screen "SP" 800x480, template "Main"
   GraphicView "Graphic view_1" at 20,61 size 347x209; Picture "clean2"
   TextField "Text field_1" at 288,5 size 156x47; Text 'Уставки'
   TextField "Text field_2" at 138,75 size 112x33; Text 'Дозация'
   TextField "Text field_12" at 28,137 size 34x23; Text 'С ='
   TextField "Text field_13" at 132,138 size 67x23; Text '% масс'
   GraphicView "Graphic view_2" at 64,133 size 66x33; Picture "input_1"
   IOField "I/O field_1" at 68,136 size 58x27; Authorization "Operator"; FormatPattern 9.99
      ProcessValue <- "Logick_DB_SP"
   GraphicView "Graphic view_5" at 368,61 size 347x209; Picture "clean2"
   TextField "Text field_21" at 436,75 size 211x33; Text 'Перемешивание'
   TextField "Text field_22" at 381,129 size 215x23; Text 'Первое перемешивание:'
   TextField "Text field_23" at 667,129 size 17x23; Text 'м'
   GraphicView "Graphic view_6" at 599,124 size 66x33; Picture "input_1"
   IOField "I/O field_3" at 603,127 size 58x27; Authorization "Operator"; FormatPattern 99
      ProcessValue <- "Logick_DB_T_M_SP_M"
   GraphicView "Graphic view_8" at 21,270 size 347x209; Picture "clean2"
   TextField "Text field_14" at 108,283 size 174x33; Text 'Реле протока'
      Visibility <- "CONFIG_Config_Use_DL"
   GraphicView "Graphic view_11" at 368,270 size 347x209; Picture "clean2"
   TextField "Text field_9" at 430,284 size 223x33; Text 'Контроль уровня'
   TextField "Text field_3" at 76,118 size 43x17; Text 'макс 1'
   TextField "Text field_4" at 71,163 size 53x17; Text 'мин 0.05'
   TextField "Text field_5" at 29,177 size 192x23; Text 'Литров на 1 дозацию:'
   TextField "Text field_6" at 29,221 size 183x23; Text 'Начало дозации при:'
   TextField "Text field_7" at 317,178 size 15x23; Text 'л'
   GraphicView "Graphic view_3" at 221,174 size 95x33; Picture "input_1"
   IOField "I/O field_2" at 227,177 size 84x27; Authorization "Operator"; FormatPattern 9999.9
      ProcessValue <- "Logick_DB_L_Per_Dos"
   TextField "Text field_26" at 291,223 size 24x23; Text '%'
   GraphicView "Graphic view_4" at 223,218 size 66x33; Picture "input_1"
   IOField "I/O field_8" at 227,221 size 58x27; Authorization "Operator"; FormatPattern 99
      ProcessValue <- "Logick_DB_L_Percent"
   TextField "Text field_27" at 231,203 size 50x17; Text 'макс 85'
   TextField "Text field_28" at 238,247 size 36x17; Text 'мин 5'
   TextField "Text field_24" at 381,163 size 168x23; Text 'Работа мешалки 1:'
   TextField "Text field_25" at 668,163 size 17x23; Text 'м'
   GraphicView "Graphic view_7" at 599,158 size 66x33; Picture "input_1"
   IOField "I/O field_9" at 603,161 size 58x27; Authorization "Operator"; FormatPattern 99
      ProcessValue <- "Logick_DB_T_M_1_SP_M"
   TextField "Text field_29" at 381,197 size 168x23; Text 'Работа мешалки 2:'
   TextField "Text field_30" at 669,197 size 17x23; Text 'м'
   GraphicView "Graphic view_14" at 599,192 size 66x33; Picture "input_1"
   IOField "I/O field_10" at 603,195 size 58x27; Authorization "Operator"; FormatPattern 99
      ProcessValue <- "Logick_DB_T_M_2_SP_M"
   TextField "Text field_31" at 381,231 size 168x23; Text 'Работа мешалки 3:'
   TextField "Text field_32" at 670,231 size 17x23; Text 'м'
   GraphicView "Graphic view_15" at 599,226 size 66x33; Picture "input_1"
   IOField "I/O field_11" at 603,229 size 58x27; Authorization "Operator"; FormatPattern 99
      ProcessValue <- "Logick_DB_T_M_3_SP_M"
   TextField "Text field_15" at 29,341 size 210x23; Text 'Отключение по датчику'
   TextField "Text field_16" at 29,376 size 197x23; Text 'Запрос на отключение'
   TextField "Text field_19" at 29,411 size 164x23; Text 'Отключение через'
   Button "Button_2" at 252,338 size 100x30; TextOff 'Text'; Authorization "Operator"; PictureList "ON_OFF"
      on Click: InvertBit("Logick_DB_DD_Stop")
      ProcessValue <- "Logick_DB_DD_Stop"
   Button "Button_3" at 252,373 size 100x30; TextOff 'Text'; Authorization "Operator"; PictureList "ON_OFF"
      on Click: InvertBit("Logick_DB_DD_REQ")
      ProcessValue <- "Logick_DB_DD_REQ"
   TextField "Text field_20" at 321,410 size 17x23; Text 'м'
   GraphicView "Graphic view_9" at 250,405 size 66x33; Picture "input_1"
   IOField "I/O field_6" at 254,408 size 58x27; Authorization "Operator"; FormatPattern 99
      ProcessValue <- "Logick_DB_T_DD_Stop_SP_M"
   TextField "Text field_10" at 374,342 size 122x23; Text 'Останов по LL'
   TextField "Text field_11" at 374,376 size 128x23; Text 'Останов по HH'
   TextField "Text field_17" at 374,411 size 197x23; Text 'Запрос на отключение'
   TextField "Text field_18" at 374,446 size 164x23; Text 'Отключение через'
   Button "Button_4" at 597,339 size 100x30; TextOff 'Text'; Authorization "Operator"; PictureList "ON_OFF"
      on Click: InvertBit("Logick_DB_LL_Stop")
      ProcessValue <- "Logick_DB_LL_Stop"
   Button "Button_5" at 597,373 size 100x30; TextOff 'Text'; Authorization "Operator"; PictureList "ON_OFF"
      on Click: InvertBit("Logick_DB_HH_Stop")
      ProcessValue <- "Logick_DB_HH_Stop"
   Button "Button_6" at 597,408 size 100x30; TextOff 'Text'; Authorization "Operator"; PictureList "ON_OFF"
      on Click: InvertBit("Logick_DB_Level_REQ")
      ProcessValue <- "Logick_DB_Level_REQ"
   TextField "Text field_33" at 666,445 size 17x23; Text 'м'
   GraphicView "Graphic view_10" at 595,440 size 66x33; Picture "input_1"
   IOField "I/O field_4" at 599,443 size 58x27; Authorization "Operator"; FormatPattern 99
      ProcessValue <- "Logick_DB_T_Level_Stop_SP_M"
   TextField "Text field_8" at 93,283 size 208x33; Text 'Низкий уровень'
      Visibility <- "CONFIG_Config_Use_DD"

screen "Calibration" 800x480, template "Main"
   GraphicView "Graphic view_1" at 20,61 size 347x209; Picture "clean2"
   TextField "Text field_1" at 256,5 size 233x47; Text 'Калибровка'
   TextField "Text field_2" at 80,75 size 225x33; Text 'Пробная дозация'
   TextField "Text field_3" at 28,161 size 33x23; Text 'q ='
   TextField "Text field_4" at 169,164 size 27x23; Text 'мл'
   TextField "Text field_5" at 28,194 size 324x23; Text 'Q = ( 60 / Тпроб ) * Тпроб * 60 / 1000'
   TextField "Text field_6" at 166,226 size 34x23; Text 'л/ч'
   TextField "Text field_7" at 28,226 size 40x23; Text 'Q ='
   TextField "Text field_12" at 28,129 size 79x23; Text 'Tпроб ='
   TextField "Text field_13" at 176,129 size 13x23; Text 'с'
   GraphicView "Graphic view_2" at 100,124 size 66x33; Picture "input_1"
   IOField "I/O field_1" at 104,127 size 58x27; Authorization "Operator"; FormatPattern 99
      ProcessValue <- "Logick_DB_T_Probe_SP_S"
   GraphicView "Graphic view_3" at 100,159 size 66x33; Picture "input_1"
   IOField "I/O field_2" at 104,162 size 58x27; Authorization "Operator"; FormatPattern 999.9
      ProcessValue <- "Logick_DB_SP_Q"
   GraphicView "Graphic view_4" at 100,221 size 66x33; Picture "input_1"
   IOField "I/O field_8" at 104,224 size 58x27; Authorization "Operator"; FormatPattern 999.9
      ProcessValue <- "Logick_DB_Q"
   GraphicView "Graphic view_5" at 368,61 size 347x209; Picture "clean2"
   TextField "Text field_21" at 487,75 size 112x33; Text 'Дозация'
   TextField "Text field_22" at 381,129 size 68x23; Text 'Tдоз ='
   TextField "Text field_23" at 556,129 size 13x23; Text 'с'
   GraphicView "Graphic view_6" at 475,124 size 66x33; Picture "input_1"
   IOField "I/O field_3" at 479,127 size 58x27; Authorization "Operator"; FormatPattern 99
      ProcessValue <- "Logick_DB_T_Dos_SP"
   TextField "Text field_24" at 546,164 size 43x23; Text 'кг/Т'
   TextField "Text field_25" at 383,164 size 71x23; Text 'Мдоз ='
   GraphicView "Graphic view_7" at 446,159 size 95x33; Picture "input_1"
   IOField "I/O field_9" at 452,162 size 84x27; Authorization "Operator"; FormatPattern 999.9999
      ProcessValue <- "Logick_DB_M_T"
   GraphicView "Graphic view_8" at 21,270 size 347x209; Picture "clean2"
   TextField "Text field_14" at 101,283 size 188x33; Text 'Концентрация'
   TextField "Text field_8" at 28,373 size 37x23; Text 'М ='
   TextField "Text field_15" at 170,376 size 42x23; Text 'кг/ч'
   TextField "Text field_16" at 28,406 size 158x23; Text 'M = ( Q * C ) / 100'
   TextField "Text field_19" at 28,341 size 34x23; Text 'С ='
   TextField "Text field_20" at 169,341 size 67x23; Text '% масс'
   GraphicView "Graphic view_9" at 100,336 size 66x33; Picture "input_1"
   IOField "I/O field_6" at 104,339 size 58x27; Authorization "Operator"; FormatPattern 999.9
      ProcessValue <- "Logick_DB_SP_C"
   GraphicView "Graphic view_10" at 100,371 size 66x33; Picture "input_1"
   IOField "I/O field_7" at 104,374 size 58x27; Authorization "Operator"; FormatPattern 999.9
      ProcessValue <- "Logick_DB_M"
   GraphicView "Graphic view_11" at 368,270 size 347x209; Picture "clean2"
   TextField "Text field_9" at 405,284 size 277x33; Text 'Поддержание уровня'
   TextField "Text field_10" at 380,376 size 72x23; Text 'Нижний'
   TextField "Text field_11" at 529,379 size 24x23; Text '%'
   TextField "Text field_17" at 380,344 size 76x23; Text 'Верхний'
   TextField "Text field_18" at 528,344 size 24x23; Text '%'
   GraphicView "Graphic view_12" at 461,339 size 66x33; Picture "input_1"
   IOField "I/O field_4" at 465,342 size 58x27; Authorization "Operator"; FormatPattern 99.9
      ProcessValue <- "AIx_DB_Level_SP_H"
   GraphicView "Graphic view_13" at 461,374 size 66x33; Picture "input_1"
   IOField "I/O field_5" at 465,377 size 58x27; Authorization "Operator"; FormatPattern 99.9
      ProcessValue <- "AIx_DB_Level_SP_L"
   Button "Button_1" at 207,126 size 144x32; TextOff 'Взять пробу'; Authorization "Operator"
      on Click: SetBit("Logick_DB_REQ_Calibration")
      Appearance <- "Logick_DB_REQ_Calibration"

screen "Monitor" 800x480, template "Main"
   Button "HmiScreenItemData_1" at 10,425 size 159x47; TextOff 'Система'; Authorization "Admin"; PictureOff "Navigates to System screens for KTP700 Basic+ PN 14.0.1.0"; PictureOn "Navigates to System screens for KTP700 Basic+ PN 14.0.1.0"
      on Release: ActivateScreen("System screens", 0)
   Button "HmiScreenItemData_2" at 195,425 size 159x47; TextOff 'Конфигурация'; Authorization "Developer"; PictureOff "Navigates to System screens for KTP700 Basic+ PN 14.0.1.0"; PictureOn "Navigates to System screens for KTP700 Basic+ PN 14.0.1.0"
      on Release: ActivateScreen("Configuration", 0)
   Button "HmiScreenItemData_3" at 380,425 size 159x47; TextOff 'Настройки'; Authorization "Admin"; PictureOff "Navigates to System screens for KTP700 Basic+ PN 14.0.1.0"; PictureOn "Navigates to System screens for KTP700 Basic+ PN 14.0.1.0"
      on Release: ActivateScreen("Settings", 0); SetTag("settings", 0)
   Button "HmiScreenItemData_4" at 565,425 size 159x47; TextOn 'О нас'; TextOff 'О нас'; PictureOn "Navigates to System screens for KTP700 Basic+ PN 14.0.1.0"; PictureOff "Navigates to System screens for KTP700 Basic+ PN 14.0.1.0"
      on Release: ActivateScreen("About", 0)
   TextField "Text field_1" at 168,4 size 424x47; Text 'Параметры установки'
   TextField "Text field_2" at 261,56 size 262x33; Text 'Состояние сигналов'
   TextField "Text field_3" at 71,92 size 189x27; Text 'Дискретные входа'
   TextField "Text field_4" at 477,92 size 205x27; Text 'Дискретные выхода'
   TextField "Text field_5" at 485,346 size 189x27; Text 'Аналоговые входа'
   TextField "Text field_6" at 43,117 size 264x23; Text 'I 0.0 - Мешалка 1 - Готовность'
   TextField "Text field_7" at 43,138 size 230x23; Text 'I 0.1 - Мешалка 1 - Работа'
   TextField "Text field_8" at 43,160 size 264x23; Text 'I 0.2 - Мешалка 2 - Готовность'
   TextField "Text field_9" at 43,181 size 230x23; Text 'I 0.3 - Мешалка 2 - Работа'
   TextField "Text field_10" at 43,203 size 264x23; Text 'I 0.4 - Мешалка 3 - Готовность'
   TextField "Text field_11" at 43,224 size 230x23; Text 'I 0.5 - Мешалка 3 - Работа'
   TextField "Text field_12" at 43,246 size 293x23; Text 'I 0.6 - Сухой дозатор - Готовность'
   TextField "Text field_13" at 43,267 size 205x23; Text 'I 0.7 - Дозатор - Работа'
   TextField "Text field_14" at 43,289 size 290x23; Text 'I 1.0 - Низкий уровень в дозаторе'
   TextField "Text field_15" at 43,310 size 250x23; Text 'I 1.1 - Вибратор - Готовность'
   TextField "Text field_16" at 43,332 size 229x23; Text 'I 1.2 - Пневмотранспортер'
   TextField "Text field_17" at 43,353 size 311x23; Text 'I 1.3 - Жидкий дозатор - Готовность'
   TextField "Text field_18" at 43,375 size 194x23; Text 'I 1.4 - Датчик протока'
   TextField "Text field_19" at 43,397 size 298x23; Text 'I 1.5 - Внешний останов / Перелив'
   Circle "Circle_1" at 10,120 size 17x17
      Appearance <- "DIx_DB_M1_FB_Ready_Signal"
   Circle "Circle_2" at 10,141 size 17x17
      Appearance <- "DIx_DB_M1_FB_Run_Signal"
   Circle "Circle_3" at 10,163 size 17x17
      Appearance <- "DIx_DB_M2_FB_Ready_Signal"
   Circle "Circle_4" at 10,184 size 17x17
      Appearance <- "DIx_DB_M2_FB_Run_Signal"
   Circle "Circle_5" at 10,206 size 17x17
      Appearance <- "DIx_DB_M3_FB_Ready_Signal"
   Circle "Circle_6" at 10,227 size 17x17
      Appearance <- "DIx_DB_M3_FB_Run_Signal"
   Circle "Circle_7" at 10,249 size 17x17
      Appearance <- "DIx_DB_DD_FB_Ready_Signal"
   Circle "Circle_8" at 10,270 size 17x17
      Appearance <- "DIx_DB_Dos_FB_Run_Signal"
   Circle "Circle_9" at 10,292 size 17x17
      Appearance <- "DIx_DB_DD_LLS_Signal"
   Circle "Circle_10" at 10,313 size 17x17
      Appearance <- "DIx_DB_Vibro_FB_Ready_Signal"
   Circle "Circle_11" at 10,335 size 17x17
      Appearance <- "DIx_DB_Transporter_Signal"
   Circle "Circle_12" at 10,356 size 17x17
      Appearance <- "DIx_DB_DL_FB_Ready_Signal"
   Circle "Circle_13" at 10,378 size 17x17
      Appearance <- "DIx_DB_Dry_Run_Signal"
   Circle "Circle_14" at 10,400 size 17x17
      Appearance <- "DIx_DB_AllBlock_Signal"
   TextField "Text field_20" at 447,117 size 232x23; Text 'Q 0.0 - Мешалка 1 - Запуск'
   TextField "Text field_21" at 447,139 size 232x23; Text 'Q 0.1 - Мешалка 2 - Запуск'
   TextField "Text field_22" at 447,160 size 232x23; Text 'Q 0.2 - Мешалка 3 - Запуск'
   TextField "Text field_23" at 447,182 size 261x23; Text 'Q 0.3 - Сухой дозатор - Запуск'
   TextField "Text field_24" at 447,203 size 218x23; Text 'Q 0.4 - Вибратор - Запуск'
   TextField "Text field_25" at 447,225 size 279x23; Text 'Q 0.5 - Жидкий дозатор - Запуск'
   TextField "Text field_26" at 447,246 size 251x23; Text 'Q 0.6 - Клапан КС1 - Открыть'
   TextField "Text field_27" at 447,268 size 221x23; Text 'Q 0.7 - Лампа - Сухой ход'
   TextField "Text field_28" at 447,289 size 258x23; Text 'Q 1.0 - Лампа - Общая авария'
   Circle "Circle_15" at 414,120 size 17x17
      Appearance <- "DOx_DB_M1_CMD_Q"
   Circle "Circle_16" at 414,142 size 17x17
      Appearance <- "DOx_DB_M2_CMD_Q"
   Circle "Circle_17" at 414,163 size 17x17
      Appearance <- "DOx_DB_M3_CMD_Q"
   Circle "Circle_18" at 414,185 size 17x17
      Appearance <- "DOx_DB_DD_CMD_Q"
   Circle "Circle_19" at 414,206 size 17x17
      Appearance <- "DOx_DB_Vibro_CMD_Q"
   Circle "Circle_20" at 414,228 size 17x17
      Appearance <- "DOx_DB_DL_CMD_Q"
   Circle "Circle_21" at 414,249 size 17x17
      Appearance <- "DOx_DB_KC1_CMD_Q"
   Circle "Circle_22" at 414,271 size 17x17
      Appearance <- "DOx_DB_LED_Dry_Run_Q"
   Circle "Circle_23" at 414,292 size 17x17
      Appearance <- "DOx_DB_LED_Alarm_Q"
   TextField "Text field_29" at 447,310 size 236x23; Text 'Q 1.1 - Лампа - Бункер пуст'
   Circle "Circle_24" at 414,313 size 17x17
      Appearance <- "DOx_DB_LED_Empty_Q"
   TextField "Text field_30" at 414,375 size 193x23; Text 'PIW 256 - Расходомер'
   TextField "Text field_31" at 414,398 size 161x23; Text 'PIW 258 - Уровень'
   IOField "I/O field_1" at 617,376 size 96x22; FormatPattern s99999
      ProcessValue <- "AIx_DB_FlowMeter_Signal"
   IOField "I/O field_2" at 617,396 size 96x22; FormatPattern s99999
      ProcessValue <- "AIx_DB_Level_Signal"

screen "Mix" 800x480, template "Main"
   Button "Button_1" at 7,5 size 96x32; TextOff 'Мешалки'; Authorization "Admin"
      on Release: ActivateScreen("Mix", 0); SetTag("settings", 1)
      Appearance <- "settings"
   Button "Button_2" at 7,52 size 96x32; TextOff 'Дозаторы'; Authorization "Admin"
      on Release: ActivateScreen("Dos", 0); SetTag("settings", 2)
      Appearance <- "settings"
   Button "Button_3" at 7,99 size 96x32; TextOff 'Клапана'; Authorization "Admin"
      on Release: ActivateScreen("Valve", 0); SetTag("settings", 3)
      Appearance <- "settings"
   Button "Button_4" at 7,146 size 96x32; TextOff 'AI'; Authorization "Admin"
      on Release: ActivateScreen("AI", 0); SetTag("settings", 4)
      Appearance <- "settings"
   Button "Button_5" at 7,193 size 96x32; TextOff 'DI'; Authorization "Admin"
      on Release: ActivateScreen("DI", 0); SetTag("settings", 5)
      Appearance <- "settings"
   Button "Button_6" at 7,240 size 96x32; TextOff 'DO'; Authorization "Admin"
      on Release: ActivateScreen("DO", 0); SetTag("settings", 6)
      Appearance <- "settings"
   Group "Group_1" at 127,146 size 416x126; Text 'Мешалка 1'; PictureList "Motor"; TextList "Hand"; Picture "z2use_3"
   Group "Group_2" at 127,285 size 416x126; Text 'Мешалка 1'; PictureList "Motor"; TextList "Hand"; Picture "z2use_3"
   Rectangle "Rectangle_1" at 127,7 size 416x126
      Appearance <- "Motors_DB_Mix_1_CMD_Sim"
   GraphicIOField "Graphic I/O field_2" at 134,43 size 43x85; PictureList "Motor"
      ProcessValue <- "Motors_DB_Mix_1_Status"
   Button "Button_7" at 213,41 size 90x22; TextOff 'Авто'; TextList "Hand"
      on Click: InvertBit("Motors_DB_Mix_1_CMD_Hand")
      Appearance <- "Motors_DB_Mix_1_CMD_Hand"
      ProcessValue <- "Motors_DB_Mix_1_CMD_Hand"
   Button "Button_8" at 258,63 size 45x22; TextOff 'Выкл'
      on Click: ResetBit("Motors_DB_Mix_1_CMD_Start_M")
   Button "Button_9" at 213,86 size 90x20; TextOff 'Сервис'
      on Click: InvertBit("Motors_DB_Mix_1_CMD_Service")
      Appearance <- "Motors_DB_Mix_1_CMD_Service"
   Button "Button_13" at 213,63 size 45x22; TextOff 'Вкл'
      on Click: SetBit("Motors_DB_Mix_1_CMD_Start_M")
      Appearance <- "Motors_DB_Mix_1_CMD_Start_M"
   TextField "Text field_13" at 133,12 size 171x26; Text 'Мешалка 1'
   TextField "Text field_15" at 310,12 size 99x18; Text 'Ожидание ОС, с'
   GraphicView "Graphic view_1" at 180,42 size 25x25; Picture "z2use_3"
      Visibility <- "Motors_DB_Mix_1_CMD_Hand"
   GraphicView "Graphic view_8" at 180,74 size 25x25; Picture "force"
      Visibility <- "Motors_DB_Mix_1_CMD_Force"
   GraphicView "Graphic view_11" at 180,103 size 25x25; Picture "service"
      Visibility <- "Motors_DB_Mix_1_CMD_Service"
   TextField "Text field_3" at 436,31 size 20x18; Text 'QF'
   TextField "Text field_10" at 436,56 size 21x18; Text 'KM'
   TextField "Text field_12" at 436,82 size 44x18; Text 'Service'
   TextField "Text field_14" at 436,108 size 41x18; Text 'Termo'
   TextField "Text field_4" at 416,10 size 120x22; Text 'Использовать:'
   Button "Button_21" at 478,32 size 60x20; TextOff 'Text'; Authorization "Operator"; PictureList "ON_OFF"
      on Click: InvertBit("Motors_DB_Mix_1_Use_QF")
      ProcessValue <- "Motors_DB_Mix_1_Use_QF"
   Button "Button_22" at 478,56 size 60x20; TextOff 'Text'; PictureList "ON_OFF"; Authorization "Operator"
      on Click: InvertBit("Motors_DB_Mix_1_Use_KM")
      ProcessValue <- "Motors_DB_Mix_1_Use_KM"
   Button "Button_24" at 478,80 size 60x20; TextOff 'Text'; PictureList "ON_OFF"; Authorization "Operator"
      on Click: InvertBit("Motors_DB_Mix_1_Use_Serivce")
      ProcessValue <- "Motors_DB_Mix_1_Use_Serivce"
   Button "Button_25" at 478,105 size 60x20; TextOff 'Text'; PictureList "ON_OFF"; Authorization "Operator"
      on Click: InvertBit("Motors_DB_Mix_1_Use_Termo")
      ProcessValue <- "Motors_DB_Mix_1_Use_Termo"
   Button "Button_26" at 416,31 size 20x20; TextOff 'Text'; Authorization "Operator"; PictureList "ok"
      ProcessValue <- "Motors_DB_Mix_1_FB_QF"
   Button "Button_27" at 416,55 size 20x20; TextOff 'Text'; PictureList "ok"; Authorization "Operator"
      ProcessValue <- "Motors_DB_Mix_1_FB_KM"
   Button "Button_29" at 416,80 size 20x20; TextOff 'Text'; PictureList "ok"; Authorization "Operator"
      ProcessValue <- "Motors_DB_Mix_1_Use_Serivce"
   Button "Button_30" at 416,105 size 20x20; TextOff 'Text'; PictureList "ok"; Authorization "Operator"
      ProcessValue <- "Motors_DB_Mix_1_FB_Termo"
   TextField "Text field_1" at 323,87 size 79x18; Text 'Наработка, ч'
   TextField "Text field_2" at 309,34 size 37x18; Text 'Старт'
   IOField "I/O field_5" at 348,32 size 30x20; FormatPattern 99
      ProcessValue <- "Motors_DB_Mix_1_Wait_On_SP"
   IOField "I/O field_12" at 348,55 size 30x20; FormatPattern 99
      ProcessValue <- "Motors_DB_Mix_1_Wait_Off_SP"
   TextField "Text field_5" at 309,55 size 32x18; Text 'Стоп'
   IOField "I/O field_13" at 378,32 size 30x20; FormatPattern 99
      ProcessValue <- "Motors_DB_Mix_1_Wait_On_Now"
   IOField "I/O field_14" at 378,55 size 30x20; FormatPattern 99
      ProcessValue <- "Motors_DB_Mix_1_Wait_Off_Now"
   IOField "I/O field_16" at 313,105 size 98x20; FormatPattern 9999999999
      ProcessValue <- "Motors_DB_Mix_1_Res_h"
   Button "Button_11" at 213,106 size 90x20; TextOff 'Force'
      on Click: InvertBit("Motors_DB_Mix_1_CMD_Force")
      Appearance <- "Motors_DB_Mix_1_CMD_Force"
   Rectangle "Rectangle_2" at 127,146 size 416x126
      Appearance <- "Motors_DB_Mix_2_CMD_Sim"
   GraphicIOField "Graphic I/O field_1" at 134,182 size 43x85; PictureList "Motor"
      ProcessValue <- "Motors_DB_Mix_2_Status"
   Button "Button_10" at 213,180 size 90x22; TextOff 'Авто'; TextList "Hand"
      on Click: InvertBit("Motors_DB_Mix_2_CMD_Hand")
      Appearance <- "Motors_DB_Mix_2_CMD_Hand"
      ProcessValue <- "Motors_DB_Mix_2_CMD_Hand"
   Button "Button_12" at 258,202 size 45x22; TextOff 'Выкл'
      on Click: ResetBit("Motors_DB_Mix_2_CMD_Start_M")
   Button "Button_14" at 213,225 size 90x20; TextOff 'Сервис'
      on Click: InvertBit("Motors_DB_Mix_2_CMD_Service")
      Appearance <- "Motors_DB_Mix_2_CMD_Service"
   Button "Button_15" at 213,202 size 45x22; TextOff 'Вкл'
      on Click: SetBit("Motors_DB_Mix_2_CMD_Start_M")
      Appearance <- "Motors_DB_Mix_2_CMD_Start_M"
   TextField "Text field_6" at 133,151 size 171x26; Text 'Мешалка 2'
   TextField "Text field_7" at 310,151 size 99x18; Text 'Ожидание ОС, с'
   GraphicView "Graphic view_2" at 180,181 size 25x25; Picture "z2use_3"
      Visibility <- "Motors_DB_Mix_2_CMD_Hand"
   GraphicView "Graphic view_3" at 180,213 size 25x25; Picture "force"
      Visibility <- "Motors_DB_Mix_2_CMD_Force"
   GraphicView "Graphic view_4" at 180,242 size 25x25; Picture "service"
      Visibility <- "Motors_DB_Mix_2_CMD_Service"
   TextField "Text field_8" at 436,170 size 20x18; Text 'QF'
   TextField "Text field_9" at 436,195 size 21x18; Text 'KM'
   TextField "Text field_11" at 436,221 size 44x18; Text 'Service'
   TextField "Text field_16" at 436,247 size 41x18; Text 'Termo'
   TextField "Text field_17" at 416,149 size 120x22; Text 'Использовать:'
   Button "Button_16" at 478,171 size 60x20; TextOff 'Text'; PictureList "ON_OFF"; Authorization "Operator"
      on Click: InvertBit("Motors_DB_Mix_2_Use_QF")
      ProcessValue <- "Motors_DB_Mix_2_Use_QF"
   Button "Button_17" at 478,195 size 60x20; TextOff 'Text'; Authorization "Operator"; PictureList "ON_OFF"
      on Click: InvertBit("Motors_DB_Mix_2_Use_KM")
      ProcessValue <- "Motors_DB_Mix_2_Use_KM"
   Button "Button_18" at 478,219 size 60x20; TextOff 'Text'; Authorization "Operator"; PictureList "ON_OFF"
      on Click: InvertBit("Motors_DB_Mix_2_Use_Serivce")
      ProcessValue <- "Motors_DB_Mix_2_Use_Serivce"
   Button "Button_19" at 478,244 size 60x20; TextOff 'Text'; Authorization "Operator"; PictureList "ON_OFF"
      on Click: InvertBit("Motors_DB_Mix_2_Use_Termo")
      ProcessValue <- "Motors_DB_Mix_2_Use_Termo"
   Button "Button_20" at 416,170 size 20x20; TextOff 'Text'; PictureList "ok"; Authorization "Operator"
      ProcessValue <- "Motors_DB_Mix_2_FB_QF"
   Button "Button_23" at 416,194 size 20x20; TextOff 'Text'; Authorization "Operator"; PictureList "ok"
      ProcessValue <- "Motors_DB_Mix_2_FB_KM"
   Button "Button_28" at 416,219 size 20x20; TextOff 'Text'; Authorization "Operator"; PictureList "ok"
      ProcessValue <- "Motors_DB_Mix_2_Use_Serivce"
   Button "Button_31" at 416,244 size 20x20; TextOff 'Text'; Authorization "Operator"; PictureList "ok"
      ProcessValue <- "Motors_DB_Mix_2_FB_Termo"
   TextField "Text field_18" at 323,226 size 79x18; Text 'Наработка, ч'
   TextField "Text field_19" at 309,173 size 37x18; Text 'Старт'
   IOField "I/O field_1" at 348,171 size 30x20; FormatPattern 99
      ProcessValue <- "Motors_DB_Mix_2_Wait_On_SP"
   IOField "I/O field_2" at 348,194 size 30x20; FormatPattern 99
      ProcessValue <- "Motors_DB_Mix_2_Wait_Off_SP"
   TextField "Text field_20" at 309,194 size 32x18; Text 'Стоп'
   IOField "I/O field_3" at 378,171 size 30x20; FormatPattern 99
      ProcessValue <- "Motors_DB_Mix_2_Wait_On_Now"
   IOField "I/O field_4" at 378,194 size 30x20; FormatPattern 99
      ProcessValue <- "Motors_DB_Mix_2_Wait_Off_Now"
   IOField "I/O field_6" at 313,244 size 98x20; FormatPattern 9999999999
      ProcessValue <- "Motors_DB_Mix_2_Res_h"
   Button "Button_32" at 213,245 size 90x20; TextOff 'Force'
      on Click: InvertBit("Motors_DB_Mix_2_CMD_Force")
      Appearance <- "Motors_DB_Mix_2_CMD_Force"
   Rectangle "Rectangle_3" at 127,285 size 416x126
      Appearance <- "Motors_DB_Mix_3_CMD_Sim"
   GraphicIOField "Graphic I/O field_3" at 134,321 size 43x85; PictureList "Motor"
      ProcessValue <- "Motors_DB_Mix_3_Status"
   Button "Button_33" at 213,319 size 90x22; TextOff 'Авто'; TextList "Hand"
      on Click: InvertBit("Motors_DB_Mix_3_CMD_Hand")
      Appearance <- "Motors_DB_Mix_3_CMD_Hand"
      ProcessValue <- "Motors_DB_Mix_3_CMD_Hand"
   Button "Button_34" at 258,341 size 45x22; TextOff 'Выкл'
      on Click: ResetBit("Motors_DB_Mix_3_CMD_Start_M")
   Button "Button_35" at 213,364 size 90x20; TextOff 'Сервис'
      on Click: InvertBit("Motors_DB_Mix_3_CMD_Service")
      Appearance <- "Motors_DB_Mix_3_CMD_Service"
   Button "Button_36" at 213,341 size 45x22; TextOff 'Вкл'
      on Click: SetBit("Motors_DB_Mix_3_CMD_Start_M")
      Appearance <- "Motors_DB_Mix_3_CMD_Start_M"
   TextField "Text field_21" at 133,290 size 171x26; Text 'Мешалка 3'
   TextField "Text field_22" at 310,290 size 99x18; Text 'Ожидание ОС, с'
   GraphicView "Graphic view_5" at 180,320 size 25x25; Picture "z2use_3"
      Visibility <- "Motors_DB_Mix_3_CMD_Hand"
   GraphicView "Graphic view_6" at 180,352 size 25x25; Picture "force"
      Visibility <- "Motors_DB_Mix_3_CMD_Force"
   GraphicView "Graphic view_7" at 180,381 size 25x25; Picture "service"
      Visibility <- "Motors_DB_Mix_3_CMD_Service"
   TextField "Text field_23" at 436,309 size 20x18; Text 'QF'
   TextField "Text field_24" at 436,334 size 21x18; Text 'KM'
   TextField "Text field_25" at 436,360 size 44x18; Text 'Service'
   TextField "Text field_26" at 436,386 size 41x18; Text 'Termo'
   TextField "Text field_27" at 416,288 size 120x22; Text 'Использовать:'
   Button "Button_37" at 478,310 size 60x20; TextOff 'Text'; PictureList "ON_OFF"; Authorization "Operator"
      on Click: InvertBit("Motors_DB_Mix_3_Use_QF")
      ProcessValue <- "Motors_DB_Mix_3_Use_QF"
   Button "Button_38" at 478,334 size 60x20; TextOff 'Text'; Authorization "Operator"; PictureList "ON_OFF"
      on Click: InvertBit("Motors_DB_Mix_3_Use_KM")
      ProcessValue <- "Motors_DB_Mix_3_Use_KM"
   Button "Button_39" at 478,358 size 60x20; TextOff 'Text'; Authorization "Operator"; PictureList "ON_OFF"
      on Click: InvertBit("Motors_DB_Mix_3_Use_Serivce")
      ProcessValue <- "Motors_DB_Mix_3_Use_Serivce"
   Button "Button_40" at 478,383 size 60x20; TextOff 'Text'; Authorization "Operator"; PictureList "ON_OFF"
      on Click: InvertBit("Motors_DB_Mix_3_Use_Termo")
      ProcessValue <- "Motors_DB_Mix_3_Use_Termo"
   Button "Button_41" at 416,309 size 20x20; TextOff 'Text'; PictureList "ok"; Authorization "Operator"
      ProcessValue <- "Motors_DB_Mix_3_FB_QF"
   Button "Button_42" at 416,333 size 20x20; TextOff 'Text'; Authorization "Operator"; PictureList "ok"
      ProcessValue <- "Motors_DB_Mix_3_FB_KM"
   Button "Button_43" at 416,358 size 20x20; TextOff 'Text'; Authorization "Operator"; PictureList "ok"
      ProcessValue <- "Motors_DB_Mix_3_Use_Serivce"
   Button "Button_44" at 416,383 size 20x20; TextOff 'Text'; Authorization "Operator"; PictureList "ok"
      ProcessValue <- "Motors_DB_Mix_3_FB_Termo"
   TextField "Text field_28" at 323,365 size 79x18; Text 'Наработка, ч'
   TextField "Text field_29" at 309,312 size 37x18; Text 'Старт'
   IOField "I/O field_7" at 348,310 size 30x20; FormatPattern 99
      ProcessValue <- "Motors_DB_Mix_3_Wait_On_SP"
   IOField "I/O field_8" at 348,333 size 30x20; FormatPattern 99
      ProcessValue <- "Motors_DB_Mix_3_Wait_Off_SP"
   TextField "Text field_30" at 309,333 size 32x18; Text 'Стоп'
   IOField "I/O field_9" at 378,310 size 30x20; FormatPattern 99
      ProcessValue <- "Motors_DB_Mix_3_Wait_On_Now"
   IOField "I/O field_10" at 378,333 size 30x20; FormatPattern 99
      ProcessValue <- "Motors_DB_Mix_3_Wait_Off_Now"
   IOField "I/O field_11" at 313,383 size 98x20; FormatPattern 9999999999
      ProcessValue <- "Motors_DB_Mix_3_Res_h"
   Button "Button_45" at 213,384 size 90x20; TextOff 'Force'
      on Click: InvertBit("Motors_DB_Mix_3_CMD_Force")
      Appearance <- "Motors_DB_Mix_3_CMD_Force"

screen "Dos" 800x480, template "Main"
   Button "Button_1" at 7,5 size 96x32; TextOff 'Мешалки'; Authorization "Admin"
      on Release: ActivateScreen("Mix", 0); SetTag("settings", 1)
      Appearance <- "settings"
   Button "Button_2" at 7,52 size 96x32; TextOff 'Дозаторы'; Authorization "Admin"
      on Release: ActivateScreen("Dos", 0); SetTag("settings", 2)
      Appearance <- "settings"
   Button "Button_3" at 7,99 size 96x32; TextOff 'Клапана'; Authorization "Admin"
      on Release: ActivateScreen("Valve", 0); SetTag("settings", 3)
      Appearance <- "settings"
   Button "Button_4" at 7,146 size 96x32; TextOff 'AI'; Authorization "Admin"
      on Release: ActivateScreen("AI", 0); SetTag("settings", 4)
      Appearance <- "settings"
   Button "Button_5" at 7,193 size 96x32; TextOff 'DI'; Authorization "Admin"
      on Release: ActivateScreen("DI", 0); SetTag("settings", 5)
      Appearance <- "settings"
   Button "Button_6" at 7,240 size 96x32; TextOff 'DO'; Authorization "Admin"
      on Release: ActivateScreen("DO", 0); SetTag("settings", 6)
      Appearance <- "settings"
   Group "Group" at 127,7 size 416x126; Text 'Мешалка 1'; PictureList "Motor"; TextList "Hand"; Picture "z2use_3"
   Group "Group_1" at 127,146 size 416x126; Text 'Мешалка 1'; PictureList "Motor"; TextList "Hand"; Picture "z2use_3"
   Group "Group_2" at 127,285 size 416x126; Text 'Мешалка 1'; PictureList "Motor"; TextList "Hand"; Picture "z2use_3"
   Rectangle "Rectangle_1" at 127,7 size 416x126
      Appearance <- "Motors_DB_DD_CMD_Sim"
   GraphicIOField "Graphic I/O field_2" at 134,43 size 43x85; PictureList "Motor"
      ProcessValue <- "Motors_DB_DD_Status"
   Button "Button_7" at 213,41 size 90x22; TextOff 'Авто'; TextList "Hand"
      on Click: InvertBit("Motors_DB_DD_CMD_Hand")
      Appearance <- "Motors_DB_DD_CMD_Hand"
      ProcessValue <- "Motors_DB_DD_CMD_Hand"
   Button "Button_8" at 258,63 size 45x22; TextOff 'Выкл'
      on Click: ResetBit("Motors_DB_DD_CMD_Start_M")
   Button "Button_9" at 213,86 size 90x20; TextOff 'Сервис'
      on Click: InvertBit("Motors_DB_DD_CMD_Service")
      Appearance <- "Motors_DB_DD_CMD_Service"
   Button "Button_13" at 213,63 size 45x22; TextOff 'Вкл'
      on Click: SetBit("Motors_DB_DD_CMD_Start_M")
      Appearance <- "Motors_DB_DD_CMD_Start_M"
   TextField "Text field_13" at 133,12 size 171x26; Text 'Сухой дозатор'
   TextField "Text field_15" at 310,12 size 99x18; Text 'Ожидание ОС, с'
   GraphicView "Graphic view_1" at 180,42 size 25x25; Picture "z2use_3"
      Visibility <- "Motors_DB_DD_CMD_Hand"
   GraphicView "Graphic view_8" at 180,74 size 25x25; Picture "force"
      Visibility <- "Motors_DB_DD_CMD_Force"
   GraphicView "Graphic view_11" at 180,103 size 25x25; Picture "service"
      Visibility <- "Motors_DB_DD_CMD_Service"
   TextField "Text field_3" at 436,31 size 20x18; Text 'QF'
   TextField "Text field_10" at 436,56 size 21x18; Text 'KM'
   TextField "Text field_12" at 436,82 size 44x18; Text 'Service'
   TextField "Text field_14" at 436,108 size 41x18; Text 'Termo'
   TextField "Text field_4" at 416,10 size 120x22; Text 'Использовать:'
   Button "Button_21" at 478,32 size 60x20; TextOff 'Text'; PictureList "ON_OFF"; Authorization "Operator"
      on Click: InvertBit("Motors_DB_DD_Use_QF")
      ProcessValue <- "Motors_DB_DD_Use_QF"
   Button "Button_22" at 478,56 size 60x20; TextOff 'Text'; Authorization "Operator"; PictureList "ON_OFF"
      on Click: InvertBit("Motors_DB_DD_Use_KM")
      ProcessValue <- "Motors_DB_DD_Use_KM"
   Button "Button_24" at 478,80 size 60x20; TextOff 'Text'; Authorization "Operator"; PictureList "ON_OFF"
      on Click: InvertBit("Motors_DB_DD_Use_Serivce")
      ProcessValue <- "Motors_DB_DD_Use_Serivce"
   Button "Button_25" at 478,105 size 60x20; TextOff 'Text'; Authorization "Operator"; PictureList "ON_OFF"
      on Click: InvertBit("Motors_DB_DD_Use_Termo")
      ProcessValue <- "Motors_DB_DD_Use_Termo"
   Button "Button_26" at 416,31 size 20x20; TextOff 'Text'; PictureList "ok"; Authorization "Operator"
      ProcessValue <- "Motors_DB_DD_FB_QF"
   Button "Button_27" at 416,55 size 20x20; TextOff 'Text'; Authorization "Operator"; PictureList "ok"
      ProcessValue <- "Motors_DB_DD_FB_KM"
   Button "Button_29" at 416,80 size 20x20; TextOff 'Text'; Authorization "Operator"; PictureList "ok"
      ProcessValue <- "Motors_DB_DD_Use_Serivce"
   Button "Button_30" at 416,105 size 20x20; TextOff 'Text'; Authorization "Operator"; PictureList "ok"
      ProcessValue <- "Motors_DB_DD_FB_Termo"
   TextField "Text field_1" at 323,87 size 79x18; Text 'Наработка, ч'
   TextField "Text field_2" at 309,34 size 37x18; Text 'Старт'
   IOField "I/O field_5" at 348,32 size 30x20; FormatPattern 99
      ProcessValue <- "Motors_DB_DD_Wait_On_SP"
   IOField "I/O field_12" at 348,55 size 30x20; FormatPattern 99
      ProcessValue <- "Motors_DB_DD_Wait_Off_SP"
   TextField "Text field_5" at 309,55 size 32x18; Text 'Стоп'
   IOField "I/O field_13" at 378,32 size 30x20; FormatPattern 99
      ProcessValue <- "Motors_DB_DD_Wait_On_Now"
   IOField "I/O field_14" at 378,55 size 30x20; FormatPattern 99
      ProcessValue <- "Motors_DB_DD_Wait_Off_Now"
   IOField "I/O field_16" at 313,105 size 98x20; FormatPattern 9999999999
      ProcessValue <- "Motors_DB_DD_Res_h"
   Button "Button_11" at 213,106 size 90x20; TextOff 'Force'
      on Click: InvertBit("Motors_DB_DD_CMD_Force")
      Appearance <- "Motors_DB_DD_CMD_Force"
   Rectangle "Rectangle_2" at 127,146 size 416x126
      Appearance <- "Motors_DB_Vibro_CMD_Sim"
   GraphicIOField "Graphic I/O field_1" at 134,182 size 43x85; PictureList "Motor"
      ProcessValue <- "Motors_DB_Vibro_Status"
   Button "Button_10" at 213,180 size 90x22; TextOff 'Авто'; TextList "Hand"
      on Click: InvertBit("Motors_DB_Vibro_CMD_Hand")
      Appearance <- "Motors_DB_Vibro_CMD_Hand"
      ProcessValue <- "Motors_DB_Vibro_CMD_Hand"
   Button "Button_12" at 258,202 size 45x22; TextOff 'Выкл'
      on Click: ResetBit("Motors_DB_Vibro_CMD_Start_M")
   Button "Button_14" at 213,225 size 90x20; TextOff 'Сервис'
      on Click: InvertBit("Motors_DB_Vibro_CMD_Service")
      Appearance <- "Motors_DB_Vibro_CMD_Service"
   Button "Button_15" at 213,202 size 45x22; TextOff 'Вкл'
      on Click: SetBit("Motors_DB_Vibro_CMD_Start_M")
      Appearance <- "Motors_DB_Vibro_CMD_Start_M"
   TextField "Text field_6" at 133,151 size 171x26; Text 'Вибратор'
   TextField "Text field_7" at 310,151 size 99x18; Text 'Ожидание ОС, с'
   GraphicView "Graphic view_2" at 180,181 size 25x25; Picture "z2use_3"
      Visibility <- "Motors_DB_Vibro_CMD_Hand"
   GraphicView "Graphic view_3" at 180,213 size 25x25; Picture "force"
      Visibility <- "Motors_DB_Vibro_CMD_Force"
   GraphicView "Graphic view_4" at 180,242 size 25x25; Picture "service"
      Visibility <- "Motors_DB_Vibro_CMD_Service"
   TextField "Text field_8" at 436,170 size 20x18; Text 'QF'
   TextField "Text field_9" at 436,195 size 21x18; Text 'KM'
   TextField "Text field_11" at 436,221 size 44x18; Text 'Service'
   TextField "Text field_16" at 436,247 size 41x18; Text 'Termo'
   TextField "Text field_17" at 416,149 size 120x22; Text 'Использовать:'
   Button "Button_16" at 478,171 size 60x20; TextOff 'Text'; Authorization "Operator"; PictureList "ON_OFF"
      on Click: InvertBit("Motors_DB_Vibro_Use_QF")
      ProcessValue <- "Motors_DB_Vibro_Use_QF"
   Button "Button_17" at 478,195 size 60x20; TextOff 'Text'; PictureList "ON_OFF"; Authorization "Operator"
      on Click: InvertBit("Motors_DB_Vibro_Use_KM")
      ProcessValue <- "Motors_DB_Vibro_Use_KM"
   Button "Button_18" at 478,219 size 60x20; TextOff 'Text'; PictureList "ON_OFF"; Authorization "Operator"
      on Click: InvertBit("Motors_DB_Vibro_Use_Serivce")
      ProcessValue <- "Motors_DB_Vibro_Use_Serivce"
   Button "Button_19" at 478,244 size 60x20; TextOff 'Text'; PictureList "ON_OFF"; Authorization "Operator"
      on Click: InvertBit("Motors_DB_Vibro_Use_Termo")
      ProcessValue <- "Motors_DB_Vibro_Use_Termo"
   Button "Button_20" at 416,170 size 20x20; TextOff 'Text'; Authorization "Operator"; PictureList "ok"
      ProcessValue <- "Motors_DB_Vibro_FB_QF"
   Button "Button_23" at 416,194 size 20x20; TextOff 'Text'; PictureList "ok"; Authorization "Operator"
      ProcessValue <- "Motors_DB_Vibro_FB_KM"
   Button "Button_28" at 416,219 size 20x20; TextOff 'Text'; PictureList "ok"; Authorization "Operator"
      ProcessValue <- "Motors_DB_Vibro_Use_Serivce"
   Button "Button_31" at 416,244 size 20x20; TextOff 'Text'; PictureList "ok"; Authorization "Operator"
      ProcessValue <- "Motors_DB_Vibro_FB_Termo"
   TextField "Text field_18" at 323,226 size 79x18; Text 'Наработка, ч'
   TextField "Text field_19" at 309,173 size 37x18; Text 'Старт'
   IOField "I/O field_1" at 348,171 size 30x20; FormatPattern 99
      ProcessValue <- "Motors_DB_Vibro_Wait_On_SP"
   IOField "I/O field_2" at 348,194 size 30x20; FormatPattern 99
      ProcessValue <- "Motors_DB_Vibro_Wait_Off_SP"
   TextField "Text field_20" at 309,194 size 32x18; Text 'Стоп'
   IOField "I/O field_3" at 378,171 size 30x20; FormatPattern 99
      ProcessValue <- "Motors_DB_Vibro_Wait_On_Now"
   IOField "I/O field_4" at 378,194 size 30x20; FormatPattern 99
      ProcessValue <- "Motors_DB_Vibro_Wait_Off_Now"
   IOField "I/O field_6" at 313,244 size 98x20; FormatPattern 9999999999
      ProcessValue <- "Motors_DB_Vibro_Res_h"
   Button "Button_32" at 213,245 size 90x20; TextOff 'Force'
      on Click: InvertBit("Motors_DB_Vibro_CMD_Force")
      Appearance <- "Motors_DB_Vibro_CMD_Force"
   Rectangle "Rectangle_3" at 127,285 size 416x126
      Appearance <- "Motors_DB_DL_CMD_Sim"
   GraphicIOField "Graphic I/O field_3" at 134,321 size 43x85; PictureList "Motor"
      ProcessValue <- "Motors_DB_DL_Status"
   Button "Button_33" at 213,319 size 90x22; TextOff 'Авто'; TextList "Hand"
      on Click: InvertBit("Motors_DB_DL_CMD_Hand")
      Appearance <- "Motors_DB_DL_CMD_Hand"
      ProcessValue <- "Motors_DB_DL_CMD_Hand"
   Button "Button_34" at 258,341 size 45x22; TextOff 'Выкл'
      on Click: ResetBit("Motors_DB_DL_CMD_Start_M")
   Button "Button_35" at 213,364 size 90x20; TextOff 'Сервис'
      on Click: InvertBit("Motors_DB_DL_CMD_Service")
      Appearance <- "Motors_DB_DL_CMD_Service"
   Button "Button_36" at 213,341 size 45x22; TextOff 'Вкл'
      on Click: SetBit("Motors_DB_DL_CMD_Start_M")
      Appearance <- "Motors_DB_DL_CMD_Start_M"
   TextField "Text field_21" at 133,290 size 171x26; Text 'Жидкий дозатор'
   TextField "Text field_22" at 310,290 size 99x18; Text 'Ожидание ОС, с'
   GraphicView "Graphic view_5" at 180,320 size 25x25; Picture "z2use_3"
      Visibility <- "Motors_DB_DL_CMD_Hand"
   GraphicView "Graphic view_6" at 180,352 size 25x25; Picture "force"
      Visibility <- "Motors_DB_DL_CMD_Force"
   GraphicView "Graphic view_7" at 180,381 size 25x25; Picture "service"
      Visibility <- "Motors_DB_DL_CMD_Service"
   TextField "Text field_23" at 436,309 size 20x18; Text 'QF'
   TextField "Text field_24" at 436,334 size 21x18; Text 'KM'
   TextField "Text field_25" at 436,360 size 44x18; Text 'Service'
   TextField "Text field_26" at 436,386 size 41x18; Text 'Termo'
   TextField "Text field_27" at 416,288 size 120x22; Text 'Использовать:'
   Button "Button_37" at 478,310 size 60x20; TextOff 'Text'; Authorization "Operator"; PictureList "ON_OFF"
      on Click: InvertBit("Motors_DB_DL_Use_QF")
      ProcessValue <- "Motors_DB_DL_Use_QF"
   Button "Button_38" at 478,334 size 60x20; TextOff 'Text'; PictureList "ON_OFF"; Authorization "Operator"
      on Click: InvertBit("Motors_DB_DL_Use_KM")
      ProcessValue <- "Motors_DB_DL_Use_KM"
   Button "Button_39" at 478,358 size 60x20; TextOff 'Text'; PictureList "ON_OFF"; Authorization "Operator"
      on Click: InvertBit("Motors_DB_DL_Use_Serivce")
      ProcessValue <- "Motors_DB_DL_Use_Serivce"
   Button "Button_40" at 478,383 size 60x20; TextOff 'Text'; PictureList "ON_OFF"; Authorization "Operator"
      on Click: InvertBit("Motors_DB_DL_Use_Termo")
      ProcessValue <- "Motors_DB_DL_Use_Termo"
   Button "Button_41" at 416,309 size 20x20; TextOff 'Text'; Authorization "Operator"; PictureList "ok"
      ProcessValue <- "Motors_DB_DL_FB_QF"
   Button "Button_42" at 416,333 size 20x20; TextOff 'Text'; PictureList "ok"; Authorization "Operator"
      ProcessValue <- "Motors_DB_DL_FB_KM"
   Button "Button_43" at 416,358 size 20x20; TextOff 'Text'; PictureList "ok"; Authorization "Operator"
      ProcessValue <- "Motors_DB_DL_Use_Serivce"
   Button "Button_44" at 416,383 size 20x20; TextOff 'Text'; PictureList "ok"; Authorization "Operator"
      ProcessValue <- "Motors_DB_DL_FB_Termo"
   TextField "Text field_28" at 323,365 size 79x18; Text 'Наработка, ч'
   TextField "Text field_29" at 309,312 size 37x18; Text 'Старт'
   IOField "I/O field_7" at 348,310 size 30x20; FormatPattern 99
      ProcessValue <- "Motors_DB_DL_Wait_On_SP"
   IOField "I/O field_8" at 348,333 size 30x20; FormatPattern 99
      ProcessValue <- "Motors_DB_DL_Wait_Off_SP"
   TextField "Text field_30" at 309,333 size 32x18; Text 'Стоп'
   IOField "I/O field_9" at 378,310 size 30x20; FormatPattern 99
      ProcessValue <- "Motors_DB_DL_Wait_On_Now"
   IOField "I/O field_10" at 378,333 size 30x20; FormatPattern 99
      ProcessValue <- "Motors_DB_DL_Wait_Off_Now"
   IOField "I/O field_11" at 313,383 size 98x20; FormatPattern 9999999999
      ProcessValue <- "Motors_DB_DL_Res_h"
   Button "Button_45" at 213,384 size 90x20; TextOff 'Force'
      on Click: InvertBit("Motors_DB_DL_CMD_Force")
      Appearance <- "Motors_DB_DL_CMD_Force"

screen "Valve" 800x480, template "Main"
   Button "Button_1" at 7,5 size 96x32; TextOff 'Мешалки'; Authorization "Admin"
      on Release: ActivateScreen("Mix", 0); SetTag("settings", 1)
      Appearance <- "settings"
   Button "Button_2" at 7,52 size 96x32; TextOff 'Дозаторы'; Authorization "Admin"
      on Release: ActivateScreen("Dos", 0); SetTag("settings", 2)
      Appearance <- "settings"
   Button "Button_3" at 7,99 size 96x32; TextOff 'Клапана'; Authorization "Admin"
      on Release: ActivateScreen("Valve", 0); SetTag("settings", 3)
      Appearance <- "settings"
   Button "Button_4" at 7,146 size 96x32; TextOff 'AI'; Authorization "Admin"
      on Release: ActivateScreen("AI", 0); SetTag("settings", 4)
      Appearance <- "settings"
   Button "Button_5" at 7,193 size 96x32; TextOff 'DI'; Authorization "Admin"
      on Release: ActivateScreen("DI", 0); SetTag("settings", 5)
      Appearance <- "settings"
   Button "Button_6" at 7,240 size 96x32; TextOff 'DO'; Authorization "Admin"
      on Release: ActivateScreen("DO", 0); SetTag("settings", 6)
      Appearance <- "settings"
   Group "Group" at 127,7 size 264x51; TextList "Hand"
   Rectangle "Rectangle_2" at 127,7 size 264x51
      Appearance <- "Micro_DB_KC1_Alarm"
   TextField "Text field_5" at 130,10 size 97x22; Text 'Клапан КС1'
   Button "Button_13" at 246,11 size 59x44; TextOff 'Авто'; TextList "Hand"
      on Click: InvertBit("Micro_DB_KC1_Hand")
      Appearance <- "Micro_DB_KC1_Hand"
      ProcessValue <- "Micro_DB_KC1_Hand"
   Button "Button_14" at 188,33 size 49x22; TextOff 'Выкл'
      on Click: ResetBit("Micro_DB_KC1_Start_M")
   Button "Button_15" at 132,33 size 47x22; TextOff 'Вкл'
      on Click: SetBit("Micro_DB_KC1_Start_M")
      Appearance <- "Micro_DB_KC1_Start_M"
   TextField "Text field_1" at 306,8 size 28x23; Text 'ОС'
   Button "Button_7" at 336,11 size 50x20; TextOff 'Text'; PictureList "ON_OFF"; Authorization "Operator"
      on Click: InvertBit("Micro_DB_KC1_No_FB")
      ProcessValue <- "Micro_DB_KC1_No_FB"
   IOField "I/O field_5" at 308,31 size 30x22; FormatPattern 99
      ProcessValue <- "Micro_DB_KC1_Wait_On_SP"
   IOField "I/O field_8" at 355,31 size 30x22; FormatPattern 99
      ProcessValue <- "Micro_DB_KC1_Wait_Off_SP"